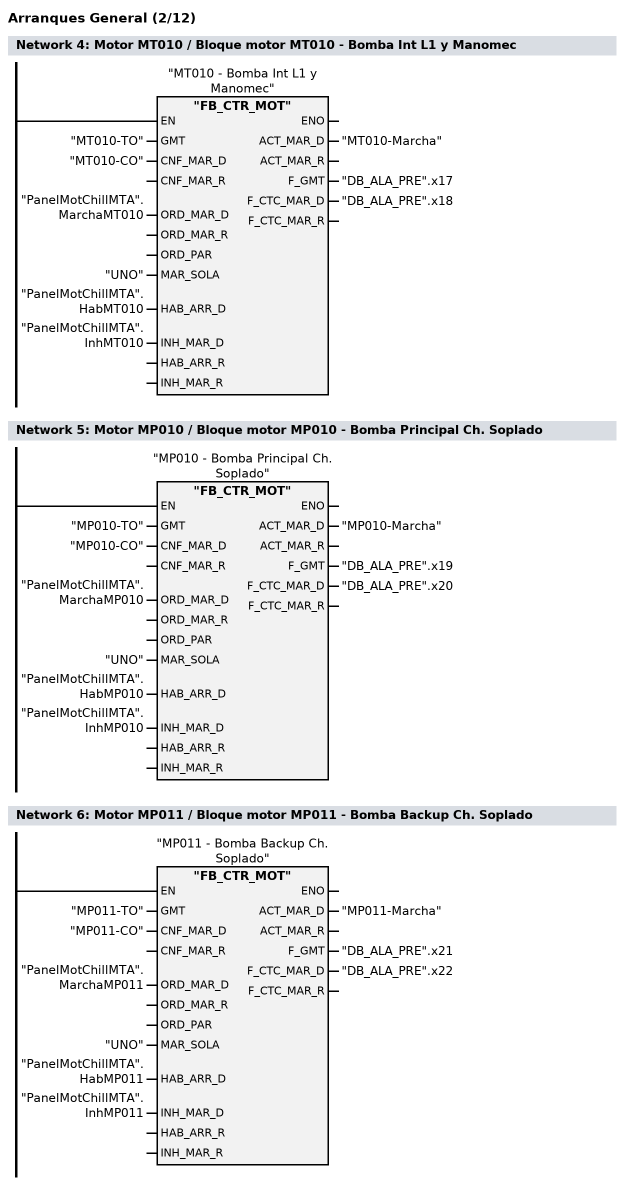
   RUNG wire#powerrail
      "MT010 - Bomba Int L1 y Manomec"(GMT := "MT010-TO", CNF_MAR_D := "MT010-CO", CNF_MAR_R :=, ORD_MAR_D := "PanelMotChillMTA".MarchaMT010, ORD_MAR_R :=, ORD_PAR :=, MAR_SOLA := "UNO", HAB_ARR_D := "PanelMotChillMTA".HabMT010, INH_MAR_D := "PanelMotChillMTA".InhMT010, HAB_ARR_R :=, INH_MAR_R :=, ACT_MAR_D => "MT010-Marcha", ACT_MAR_R =>, F_GMT => "DB_ALA_PRE".x17, F_CTC_MAR_D => "DB_ALA_PRE".x18, F_CTC_MAR_R =>)
   END_RUNG
   // the same network as SCL:
   "MT010 - Bomba Int L1 y Manomec"(GMT := "MT010-TO",   // "FB_CTR_MOT"
                           CNF_MAR_D := "MT010-CO",
                           ORD_MAR_D := "PanelMotChillMTA".MarchaMT010,
                           MAR_SOLA := "UNO",
                           HAB_ARR_D := "PanelMotChillMTA".HabMT010,
                           INH_MAR_D := "PanelMotChillMTA".InhMT010,
                           ACT_MAR_D => "MT010-Marcha",
                           F_GMT => "DB_ALA_PRE".x17,
                           F_CTC_MAR_D => "DB_ALA_PRE".x18);
END_REGION

REGION Network 5: Motor MP010 / Bloque motor MP010 - Bomba Principal Ch. Soplado
   RUNG wire#powerrail
      "MP010 - Bomba Principal Ch. Soplado"(GMT := "MP010-TO", CNF_MAR_D := "MP010-CO", CNF_MAR_R :=, ORD_MAR_D := "PanelMotChillMTA".MarchaMP010, ORD_MAR_R :=, ORD_PAR :=, MAR_SOLA := "UNO", HAB_ARR_D := "PanelMotChillMTA".HabMP010, INH_MAR_D := "PanelMotChillMTA".InhMP010, HAB_ARR_R :=, INH_MAR_R :=, ACT_MAR_D => "MP010-Marcha", ACT_MAR_R =>, F_GMT => "DB_ALA_PRE".x19, F_CTC_MAR_D => "DB_ALA_PRE".x20, F_CTC_MAR_R =>)
   END_RUNG
   // the same network as SCL:
   "MP010 - Bomba Principal Ch. Soplado"(GMT := "MP010-TO",   // "FB_CTR_MOT"
                           CNF_MAR_D := "MP010-CO",
                           ORD_MAR_D := "PanelMotChillMTA".MarchaMP010,
                           MAR_SOLA := "UNO",
                           HAB_ARR_D := "PanelMotChillMTA".HabMP010,
                           INH_MAR_D := "PanelMotChillMTA".InhMP010,
                           ACT_MAR_D => "MP010-Marcha",
                           F_GMT => "DB_ALA_PRE".x19,
                           F_CTC_MAR_D => "DB_ALA_PRE".x20);
END_REGION

REGION Network 6: Motor MP011 / Bloque motor MP011 - Bomba Backup Ch. Soplado
   RUNG wire#powerrail
      "MP011 - Bomba Backup Ch. Soplado"(GMT := "MP011-TO", CNF_MAR_D := "MP011-CO", CNF_MAR_R :=, ORD_MAR_D := "PanelMotChillMTA".MarchaMP011, ORD_MAR_R :=, ORD_PAR :=, MAR_SOLA := "UNO", HAB_ARR_D := "PanelMotChillMTA".HabMP011, INH_MAR_D := "PanelMotChillMTA".InhMP011, HAB_ARR_R :=, INH_MAR_R :=, ACT_MAR_D => "MP011-Marcha", ACT_MAR_R =>, F_GMT => "DB_ALA_PRE".x21, F_CTC_MAR_D => "DB_ALA_PRE".x22, F_CTC_MAR_R =>)
   END_RUNG
   // the same network as SCL:
   "MP011 - Bomba Backup Ch. Soplado"(GMT := "MP011-TO",   // "FB_CTR_MOT"
                           CNF_MAR_D := "MP011-CO",
                           ORD_MAR_D := "PanelMotChillMTA".MarchaMP011,
                           MAR_SOLA := "UNO",
                           HAB_ARR_D := "PanelMotChillMTA".HabMP011,
                           INH_MAR_D := "PanelMotChillMTA".InhMP011,
                           ACT_MAR_D => "MP011-Marcha",
                           F_GMT => "DB_ALA_PRE".x21,
                           F_CTC_MAR_D => "DB_ALA_PRE".x22);
END_REGION

REGION Network 7: Motor MP012 / Bloque motor MP012 - Bomba Principal Ch. Envasado
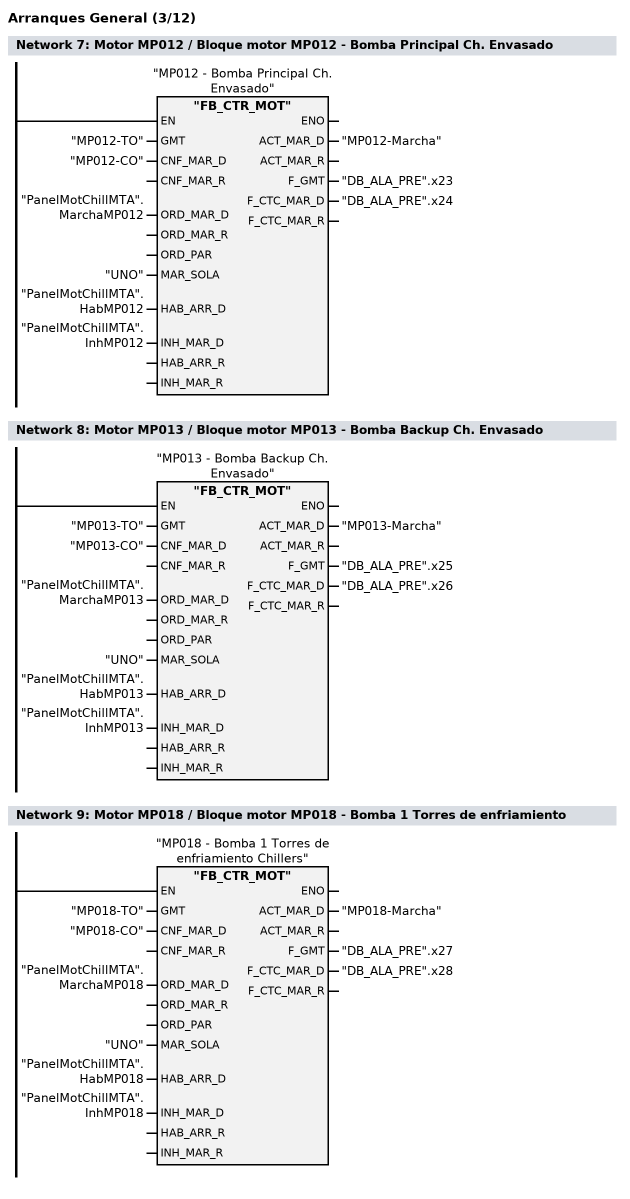
   RUNG wire#powerrail
      "MP012 - Bomba Principal Ch. Envasado"(GMT := "MP012-TO", CNF_MAR_D := "MP012-CO", CNF_MAR_R :=, ORD_MAR_D := "PanelMotChillMTA".MarchaMP012, ORD_MAR_R :=, ORD_PAR :=, MAR_SOLA := "UNO", HAB_ARR_D := "PanelMotChillMTA".HabMP012, INH_MAR_D := "PanelMotChillMTA".InhMP012, HAB_ARR_R :=, INH_MAR_R :=, ACT_MAR_D => "MP012-Marcha", ACT_MAR_R =>, F_GMT => "DB_ALA_PRE".x23, F_CTC_MAR_D => "DB_ALA_PRE".x24, F_CTC_MAR_R =>)
   END_RUNG
   // the same network as SCL:
   "MP012 - Bomba Principal Ch. Envasado"(GMT := "MP012-TO",   // "FB_CTR_MOT"
                           CNF_MAR_D := "MP012-CO",
                           ORD_MAR_D := "PanelMotChillMTA".MarchaMP012,
                           MAR_SOLA := "UNO",
                           HAB_ARR_D := "PanelMotChillMTA".HabMP012,
                           INH_MAR_D := "PanelMotChillMTA".InhMP012,
                           ACT_MAR_D => "MP012-Marcha",
                           F_GMT => "DB_ALA_PRE".x23,
                           F_CTC_MAR_D => "DB_ALA_PRE".x24);
END_REGION

REGION Network 8: Motor MP013 / Bloque motor MP013 - Bomba Backup Ch. Envasado
   RUNG wire#powerrail
      "MP013 - Bomba Backup Ch. Envasado"(GMT := "MP013-TO", CNF_MAR_D := "MP013-CO", CNF_MAR_R :=, ORD_MAR_D := "PanelMotChillMTA".MarchaMP013, ORD_MAR_R :=, ORD_PAR :=, MAR_SOLA := "UNO", HAB_ARR_D := "PanelMotChillMTA".HabMP013, INH_MAR_D := "PanelMotChillMTA".InhMP013, HAB_ARR_R :=, INH_MAR_R :=, ACT_MAR_D => "MP013-Marcha", ACT_MAR_R =>, F_GMT => "DB_ALA_PRE".x25, F_CTC_MAR_D => "DB_ALA_PRE".x26, F_CTC_MAR_R =>)
   END_RUNG
   // the same network as SCL:
   "MP013 - Bomba Backup Ch. Envasado"(GMT := "MP013-TO",   // "FB_CTR_MOT"
                           CNF_MAR_D := "MP013-CO",
                           ORD_MAR_D := "PanelMotChillMTA".MarchaMP013,
                           MAR_SOLA := "UNO",
                           HAB_ARR_D := "PanelMotChillMTA".HabMP013,
                           INH_MAR_D := "PanelMotChillMTA".InhMP013,
                           ACT_MAR_D => "MP013-Marcha",
                           F_GMT => "DB_ALA_PRE".x25,
                           F_CTC_MAR_D => "DB_ALA_PRE".x26);
END_REGION

REGION Network 9: Motor MP018 / Bloque motor MP018 - Bomba 1 Torres de enfriamiento
   RUNG wire#powerrail
      "MP018 - Bomba 1 Torres de enfriamiento Chillers"(GMT := "MP018-TO", CNF_MAR_D := "MP018-CO", CNF_MAR_R :=, ORD_MAR_D := "PanelMotChillMTA".MarchaMP018, ORD_MAR_R :=, ORD_PAR :=, MAR_SOLA := "UNO", HAB_ARR_D := "PanelMotChillMTA".HabMP018, INH_MAR_D := "PanelMotChillMTA".InhMP018, HAB_ARR_R :=, INH_MAR_R :=, ACT_MAR_D => "MP018-Marcha", ACT_MAR_R =>, F_GMT => "DB_ALA_PRE".x27, F_CTC_MAR_D => "DB_ALA_PRE".x28, F_CTC_MAR_R =>)
   END_RUNG
   // the same network as SCL:
   "MP018 - Bomba 1 Torres de enfriamiento Chillers"(GMT := "MP018-TO",   // "FB_CTR_MOT"
                           CNF_MAR_D := "MP018-CO",
                           ORD_MAR_D := "PanelMotChillMTA".MarchaMP018,
                           MAR_SOLA := "UNO",
                           HAB_ARR_D := "PanelMotChillMTA".HabMP018,
                           INH_MAR_D := "PanelMotChillMTA".InhMP018,
                           ACT_MAR_D => "MP018-Marcha",
                           F_GMT => "DB_ALA_PRE".x27,
                           F_CTC_MAR_D => "DB_ALA_PRE".x28);
END_REGION

REGION Network 10: Motor MP019 / Bloque motor MP019 - Bomba 2 Torres de enfriamiento
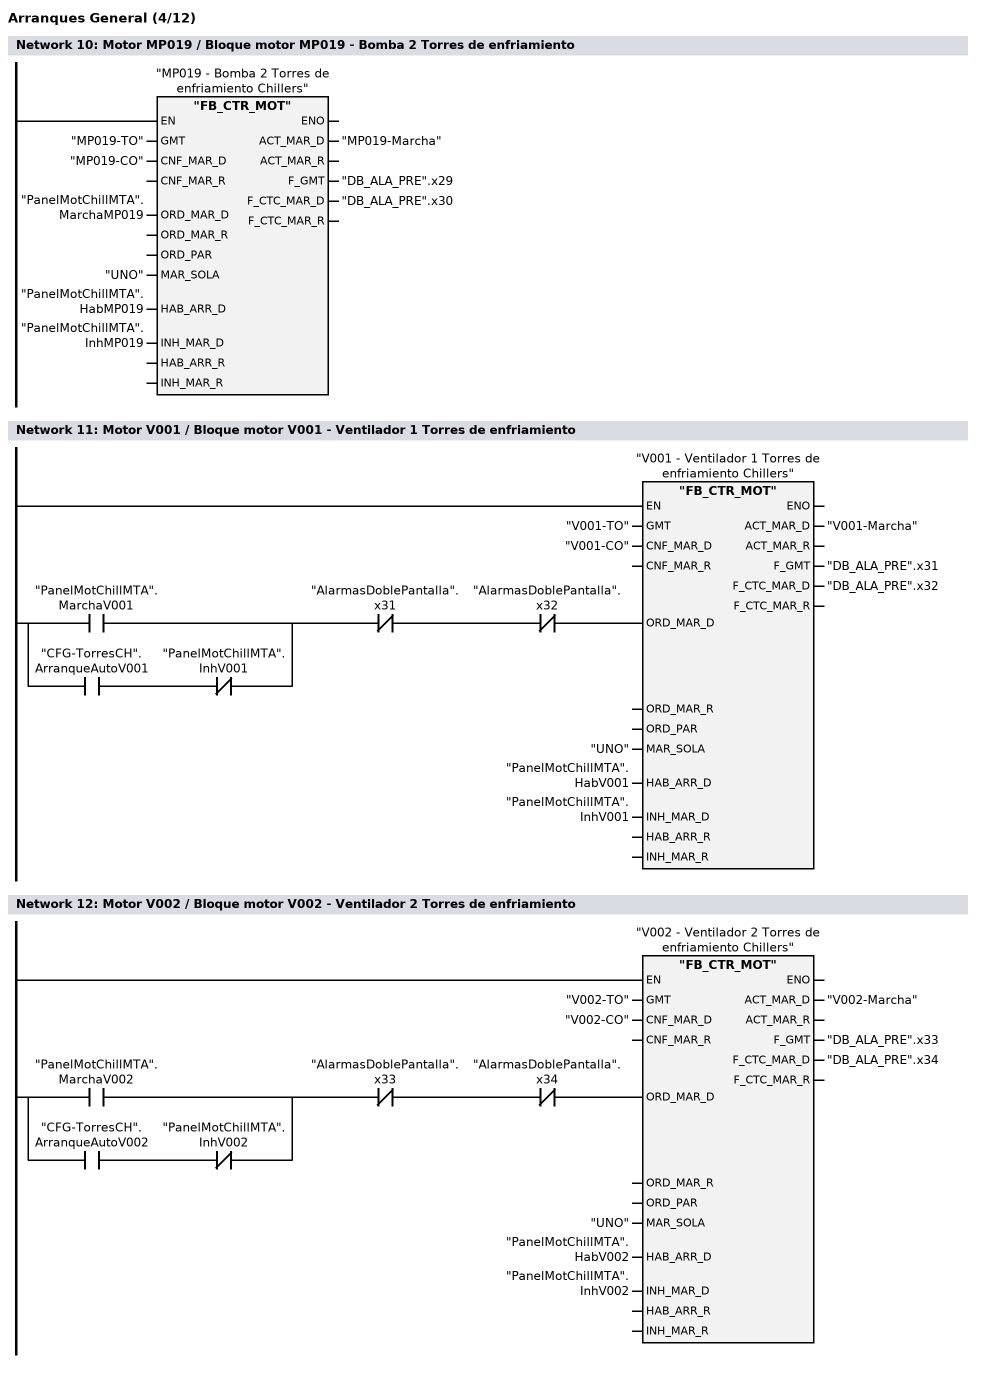
   RUNG wire#powerrail
      "MP019 - Bomba 2 Torres de enfriamiento Chillers"(GMT := "MP019-TO", CNF_MAR_D := "MP019-CO", CNF_MAR_R :=, ORD_MAR_D := "PanelMotChillMTA".MarchaMP019, ORD_MAR_R :=, ORD_PAR :=, MAR_SOLA := "UNO", HAB_ARR_D := "PanelMotChillMTA".HabMP019, INH_MAR_D := "PanelMotChillMTA".InhMP019, HAB_ARR_R :=, INH_MAR_R :=, ACT_MAR_D => "MP019-Marcha", ACT_MAR_R =>, F_GMT => "DB_ALA_PRE".x29, F_CTC_MAR_D => "DB_ALA_PRE".x30, F_CTC_MAR_R =>)
   END_RUNG
   // the same network as SCL:
   "MP019 - Bomba 2 Torres de enfriamiento Chillers"(GMT := "MP019-TO",   // "FB_CTR_MOT"
                           CNF_MAR_D := "MP019-CO",
                           ORD_MAR_D := "PanelMotChillMTA".MarchaMP019,
                           MAR_SOLA := "UNO",
                           HAB_ARR_D := "PanelMotChillMTA".HabMP019,
                           INH_MAR_D := "PanelMotChillMTA".InhMP019,
                           ACT_MAR_D => "MP019-Marcha",
                           F_GMT => "DB_ALA_PRE".x29,
                           F_CTC_MAR_D => "DB_ALA_PRE".x30);
END_REGION

REGION Network 11: Motor V001 / Bloque motor V001 - Ventilador 1 Torres de enfriamiento
   RUNG wire#powerrail
      "V001 - Ventilador 1 Torres de enfriamiento Chillers"(ORD_MAR_D := wire#w2, GMT := "V001-TO", CNF_MAR_D := "V001-CO", CNF_MAR_R :=, ORD_MAR_R :=, ORD_PAR :=, MAR_SOLA := "UNO", HAB_ARR_D := "PanelMotChillMTA".HabV001, INH_MAR_D := "PanelMotChillMTA".InhV001, HAB_ARR_R :=, INH_MAR_R :=, ACT_MAR_D => "V001-Marcha", ACT_MAR_R =>, F_GMT => "DB_ALA_PRE".x31, F_CTC_MAR_D => "DB_ALA_PRE".x32, F_CTC_MAR_R =>)
   END_RUNG
   RUNG wire#powerrail
      Contact( "PanelMotChillMTA".MarchaV001 )
      wire#w1
      I_Contact( "AlarmasDoblePantalla".x31 )
      I_Contact( "AlarmasDoblePantalla".x32 )
   END_RUNG wire#w2
   RUNG wire#powerrail
      Contact( "CFG-TorresCH".ArranqueAutoV001 )
      I_Contact( "PanelMotChillMTA".InhV001 )
   END_RUNG wire#w1
   // the same network as SCL:
   "V001 - Ventilador 1 Torres de enfriamiento Chillers"(GMT := "V001-TO",   // "FB_CTR_MOT"
                           CNF_MAR_D := "V001-CO",
                           ORD_MAR_D := ("PanelMotChillMTA".MarchaV001 OR ("CFG-TorresCH".ArranqueAutoV001 AND NOT "PanelMotChillMTA".InhV001)) AND NOT "AlarmasDoblePantalla".x31 AND NOT "AlarmasDoblePantalla".x32,
                           MAR_SOLA := "UNO",
                           HAB_ARR_D := "PanelMotChillMTA".HabV001,
                           INH_MAR_D := "PanelMotChillMTA".InhV001,
                           ACT_MAR_D => "V001-Marcha",
                           F_GMT => "DB_ALA_PRE".x31,
                           F_CTC_MAR_D => "DB_ALA_PRE".x32);
END_REGION

REGION Network 12: Motor V002 / Bloque motor V002 - Ventilador 2 Torres de enfriamiento
   RUNG wire#powerrail
      "V002 - Ventilador 2 Torres de enfriamiento Chillers"(ORD_MAR_D := wire#w2, GMT := "V002-TO", CNF_MAR_D := "V002-CO", CNF_MAR_R :=, ORD_MAR_R :=, ORD_PAR :=, MAR_SOLA := "UNO", HAB_ARR_D := "PanelMotChillMTA".HabV002, INH_MAR_D := "PanelMotChillMTA".InhV002, HAB_ARR_R :=, INH_MAR_R :=, ACT_MAR_D => "V002-Marcha", ACT_MAR_R =>, F_GMT => "DB_ALA_PRE".x33, F_CTC_MAR_D => "DB_ALA_PRE".x34, F_CTC_MAR_R =>)
   END_RUNG
   RUNG wire#powerrail
      Contact( "PanelMotChillMTA".MarchaV002 )
      wire#w1
      I_Contact( "AlarmasDoblePantalla".x33 )
      I_Contact( "AlarmasDoblePantalla".x34 )
   END_RUNG wire#w2
   RUNG wire#powerrail
      Contact( "CFG-TorresCH".ArranqueAutoV002 )
      I_Contact( "PanelMotChillMTA".InhV002 )
   END_RUNG wire#w1
   // the same network as SCL:
   "V002 - Ventilador 2 Torres de enfriamiento Chillers"(GMT := "V002-TO",   // "FB_CTR_MOT"
                           CNF_MAR_D := "V002-CO",
                           ORD_MAR_D := ("PanelMotChillMTA".MarchaV002 OR ("CFG-TorresCH".ArranqueAutoV002 AND NOT "PanelMotChillMTA".InhV002)) AND NOT "AlarmasDoblePantalla".x33 AND NOT "AlarmasDoblePantalla".x34,
                           MAR_SOLA := "UNO",
                           HAB_ARR_D := "PanelMotChillMTA".HabV002,
                           INH_MAR_D := "PanelMotChillMTA".InhV002,
                           ACT_MAR_D => "V002-Marcha",
                           F_GMT => "DB_ALA_PRE".x33,
                           F_CTC_MAR_D => "DB_ALA_PRE".x34);
END_REGION

REGION Network 13: Motor V003 / Bloque motor V003 - Ventilador 3 Torres de enfriamiento
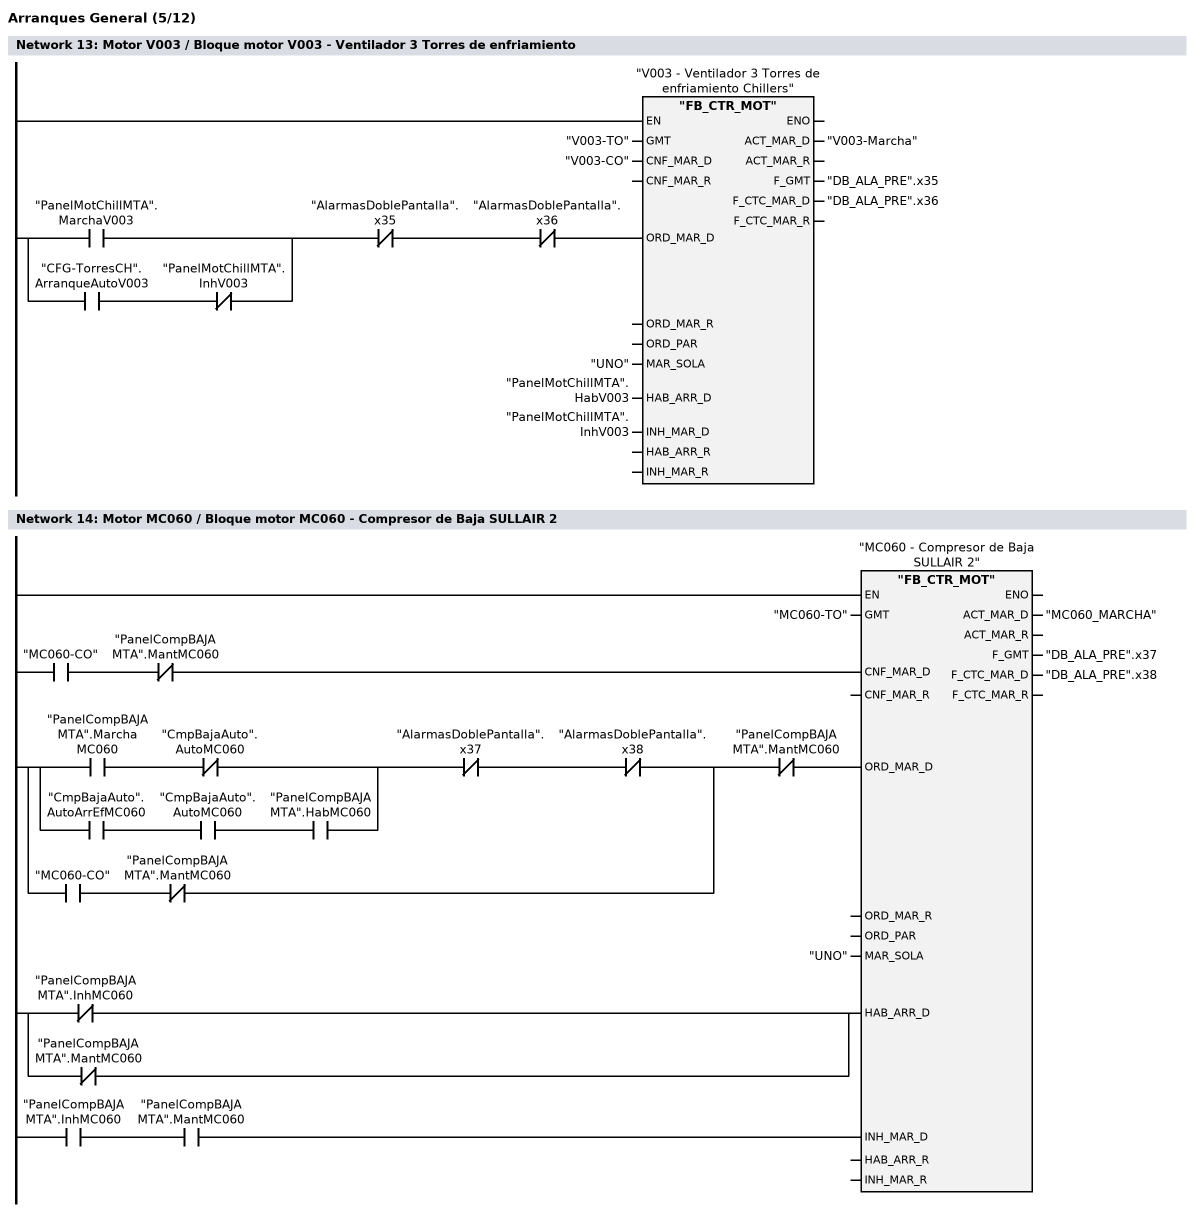
   RUNG wire#powerrail
      "V003 - Ventilador 3 Torres de enfriamiento Chillers"(ORD_MAR_D := wire#w2, GMT := "V003-TO", CNF_MAR_D := "V003-CO", CNF_MAR_R :=, ORD_MAR_R :=, ORD_PAR :=, MAR_SOLA := "UNO", HAB_ARR_D := "PanelMotChillMTA".HabV003, INH_MAR_D := "PanelMotChillMTA".InhV003, HAB_ARR_R :=, INH_MAR_R :=, ACT_MAR_D => "V003-Marcha", ACT_MAR_R =>, F_GMT => "DB_ALA_PRE".x35, F_CTC_MAR_D => "DB_ALA_PRE".x36, F_CTC_MAR_R =>)
   END_RUNG
   RUNG wire#powerrail
      Contact( "PanelMotChillMTA".MarchaV003 )
      wire#w1
      I_Contact( "AlarmasDoblePantalla".x35 )
      I_Contact( "AlarmasDoblePantalla".x36 )
   END_RUNG wire#w2
   RUNG wire#powerrail
      Contact( "CFG-TorresCH".ArranqueAutoV003 )
      I_Contact( "PanelMotChillMTA".InhV003 )
   END_RUNG wire#w1
   // the same network as SCL:
   "V003 - Ventilador 3 Torres de enfriamiento Chillers"(GMT := "V003-TO",   // "FB_CTR_MOT"
                           CNF_MAR_D := "V003-CO",
                           ORD_MAR_D := ("PanelMotChillMTA".MarchaV003 OR ("CFG-TorresCH".ArranqueAutoV003 AND NOT "PanelMotChillMTA".InhV003)) AND NOT "AlarmasDoblePantalla".x35 AND NOT "AlarmasDoblePantalla".x36,
                           MAR_SOLA := "UNO",
                           HAB_ARR_D := "PanelMotChillMTA".HabV003,
                           INH_MAR_D := "PanelMotChillMTA".InhV003,
                           ACT_MAR_D => "V003-Marcha",
                           F_GMT => "DB_ALA_PRE".x35,
                           F_CTC_MAR_D => "DB_ALA_PRE".x36);
END_REGION

REGION Network 14: Motor MC060 / Bloque motor MC060 - Compresor de Baja SULLAIR 2
   RUNG wire#powerrail
      "MC060 - Compresor de Baja SULLAIR 2"(CNF_MAR_D := wire#w1, ORD_MAR_D := wire#w4, HAB_ARR_D := wire#w5, INH_MAR_D := wire#w6, GMT := "MC060-TO", CNF_MAR_R :=, ORD_MAR_R :=, ORD_PAR :=, MAR_SOLA := "UNO", HAB_ARR_R :=, INH_MAR_R :=, ACT_MAR_D => "MC060_MARCHA", ACT_MAR_R =>, F_GMT => "DB_ALA_PRE".x37, F_CTC_MAR_D => "DB_ALA_PRE".x38, F_CTC_MAR_R =>)
   END_RUNG
   RUNG wire#powerrail
      Contact( "MC060-CO" )
      I_Contact( "PanelCompBAJA MTA".MantMC060 )
   END_RUNG wire#w1
   RUNG wire#powerrail
      Contact( "PanelCompBAJA MTA".MarchaMC060 )
      I_Contact( "CmpBajaAuto".AutoMC060 )
      wire#w2
      I_Contact( "AlarmasDoblePantalla".x37 )
      I_Contact( "AlarmasDoblePantalla".x38 )
      wire#w3
      I_Contact( "PanelCompBAJA MTA".MantMC060 )
   END_RUNG wire#w4
   RUNG wire#powerrail
      Contact( "CmpBajaAuto".AutoArrEfMC060 )
      Contact( "CmpBajaAuto".AutoMC060 )
      Contact( "PanelCompBAJA MTA".HabMC060 )
   END_RUNG wire#w2
   RUNG wire#powerrail
      Contact( "MC060-CO" )
      I_Contact( "PanelCompBAJA MTA".MantMC060 )
   END_RUNG wire#w3
   RUNG wire#powerrail
      I_Contact( "PanelCompBAJA MTA".InhMC060 )
   END_RUNG wire#w5
   RUNG wire#powerrail
      I_Contact( "PanelCompBAJA MTA".MantMC060 )
   END_RUNG wire#w5
   RUNG wire#powerrail
      Contact( "PanelCompBAJA MTA".InhMC060 )
      Contact( "PanelCompBAJA MTA".MantMC060 )
   END_RUNG wire#w6
   // the same network as SCL:
   "MC060 - Compresor de Baja SULLAIR 2"(GMT := "MC060-TO",   // "FB_CTR_MOT"
                           CNF_MAR_D := "MC060-CO" AND NOT "PanelCompBAJA MTA".MantMC060,
                           ORD_MAR_D := (((("PanelCompBAJA MTA".MarchaMC060 AND NOT "CmpBajaAuto".AutoMC060) OR ("CmpBajaAuto".AutoArrEfMC060 AND "CmpBajaAuto".AutoMC060 AND "PanelCompBAJA MTA".HabMC060)) AND NOT "AlarmasDoblePantalla".x37 AND NOT "AlarmasDoblePantalla".x38) OR ("MC060-CO" AND NOT "PanelCompBAJA MTA".MantMC060)) AND NOT "PanelCompBAJA MTA".MantMC060,
                           MAR_SOLA := "UNO",
                           HAB_ARR_D := NOT "PanelCompBAJA MTA".InhMC060 OR NOT "PanelCompBAJA MTA".MantMC060,
                           INH_MAR_D := "PanelCompBAJA MTA".InhMC060 AND "PanelCompBAJA MTA".MantMC060,
                           ACT_MAR_D => "MC060_MARCHA",
                           F_GMT => "DB_ALA_PRE".x37,
                           F_CTC_MAR_D => "DB_ALA_PRE".x38);
END_REGION

REGION Network 15
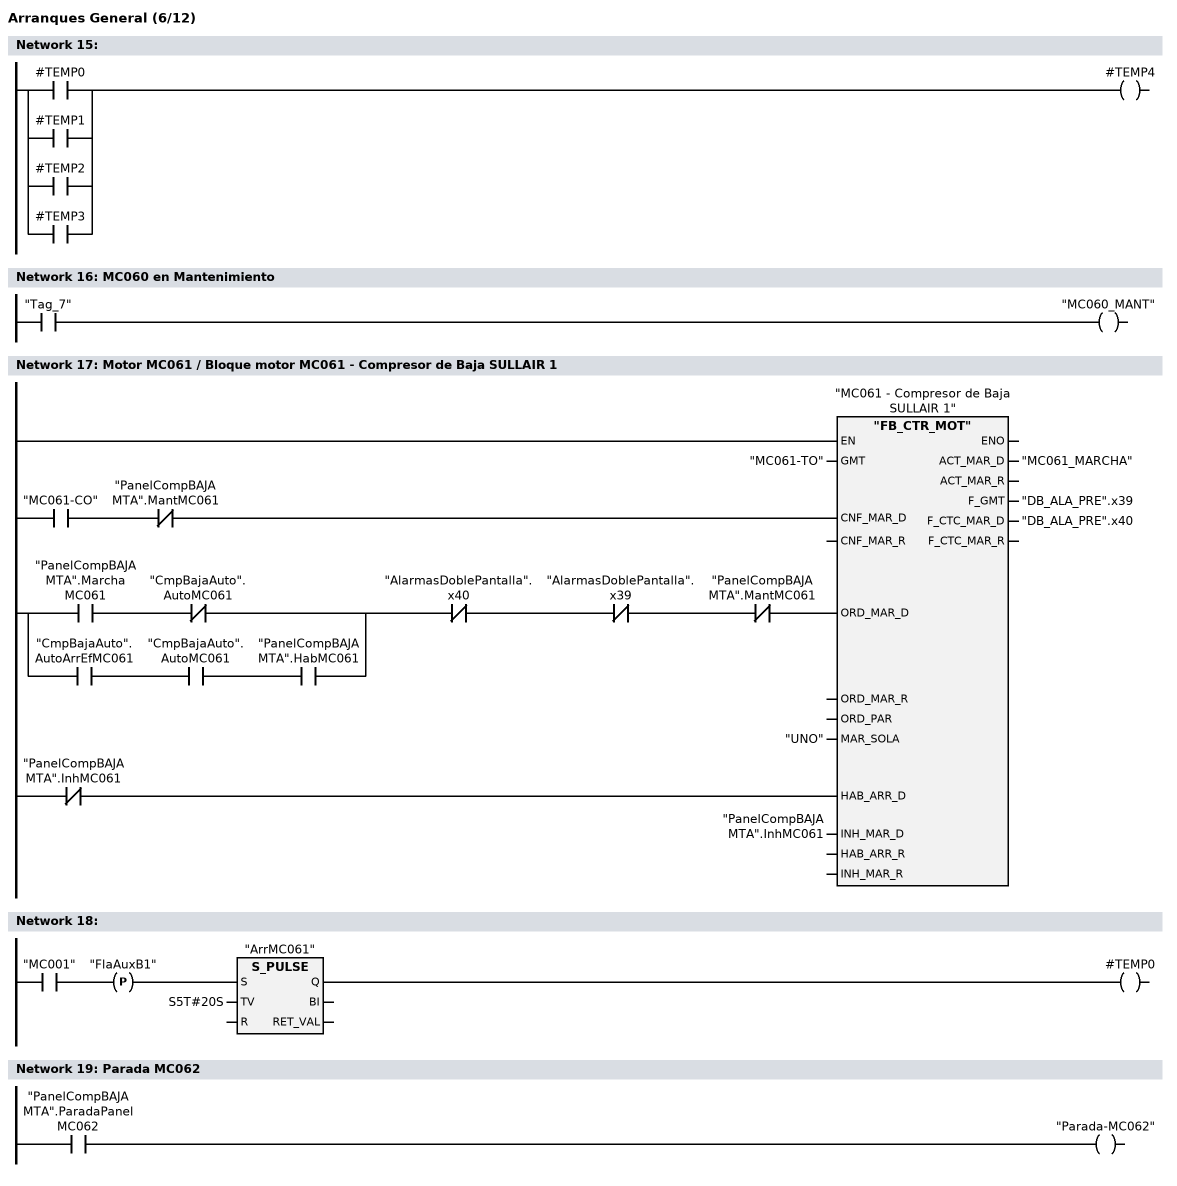
   RUNG wire#powerrail
      Contact( #TEMP0 )
      wire#w1
      Coil( #TEMP4 )
   END_RUNG
   RUNG wire#powerrail
      Contact( #TEMP1 )
   END_RUNG wire#w1
   RUNG wire#powerrail
      Contact( #TEMP2 )
   END_RUNG wire#w1
   RUNG wire#powerrail
      Contact( #TEMP3 )
   END_RUNG wire#w1
   // the same network as SCL:
   #TEMP4 := #TEMP0 OR #TEMP1 OR #TEMP2 OR #TEMP3;
END_REGION

REGION Network 16: MC060 en Mantenimiento
   RUNG wire#powerrail
      Contact( "Tag_7" )
      Coil( "MC060_MANT" )
   END_RUNG
   // the same network as SCL:
   "MC060_MANT" := "Tag_7";
END_REGION

REGION Network 17: Motor MC061 / Bloque motor MC061 - Compresor de Baja SULLAIR 1
   RUNG wire#powerrail
      "MC061 - Compresor de Baja SULLAIR 1"(CNF_MAR_D := wire#w1, ORD_MAR_D := wire#w3, HAB_ARR_D := wire#w4, GMT := "MC061-TO", CNF_MAR_R :=, ORD_MAR_R :=, ORD_PAR :=, MAR_SOLA := "UNO", INH_MAR_D := "PanelCompBAJA MTA".InhMC061, HAB_ARR_R :=, INH_MAR_R :=, ACT_MAR_D => "MC061_MARCHA", ACT_MAR_R =>, F_GMT => "DB_ALA_PRE".x39, F_CTC_MAR_D => "DB_ALA_PRE".x40, F_CTC_MAR_R =>)
   END_RUNG
   RUNG wire#powerrail
      Contact( "MC061-CO" )
      I_Contact( "PanelCompBAJA MTA".MantMC061 )
   END_RUNG wire#w1
   RUNG wire#powerrail
      Contact( "PanelCompBAJA MTA".MarchaMC061 )
      I_Contact( "CmpBajaAuto".AutoMC061 )
      wire#w2
      I_Contact( "AlarmasDoblePantalla".x40 )
      I_Contact( "AlarmasDoblePantalla".x39 )
      I_Contact( "PanelCompBAJA MTA".MantMC061 )
   END_RUNG wire#w3
   RUNG wire#powerrail
      Contact( "CmpBajaAuto".AutoArrEfMC061 )
      Contact( "CmpBajaAuto".AutoMC061 )
      Contact( "PanelCompBAJA MTA".HabMC061 )
   END_RUNG wire#w2
   RUNG wire#powerrail
      I_Contact( "PanelCompBAJA MTA".InhMC061 )
   END_RUNG wire#w4
   // the same network as SCL:
   "MC061 - Compresor de Baja SULLAIR 1"(GMT := "MC061-TO",   // "FB_CTR_MOT"
                           CNF_MAR_D := "MC061-CO" AND NOT "PanelCompBAJA MTA".MantMC061,
                           ORD_MAR_D := (("PanelCompBAJA MTA".MarchaMC061 AND NOT "CmpBajaAuto".AutoMC061) OR ("CmpBajaAuto".AutoArrEfMC061 AND "CmpBajaAuto".AutoMC061 AND "PanelCompBAJA MTA".HabMC061)) AND NOT "AlarmasDoblePantalla".x40 AND NOT "AlarmasDoblePantalla".x39 AND NOT "PanelCompBAJA MTA".MantMC061,
                           MAR_SOLA := "UNO",
                           HAB_ARR_D := NOT "PanelCompBAJA MTA".InhMC061,
                           INH_MAR_D := "PanelCompBAJA MTA".InhMC061,
                           ACT_MAR_D => "MC061_MARCHA",
                           F_GMT => "DB_ALA_PRE".x39,
                           F_CTC_MAR_D => "DB_ALA_PRE".x40);
END_REGION

REGION Network 18
   RUNG wire#powerrail
      Contact( "MC001" )
      P_Trig( "FlaAuxB1" )
      S_PULSE(T_NO := "ArrMC061", TV := S5T#20S, R :=, BI =>, RET_VAL =>)
      Coil( #TEMP0 )
   END_RUNG
   // the same network as SCL:
   #_w1 := "MC001" AND NOT "FlaAuxB1";   // rising edge
   "FlaAuxB1" := "MC001";
   #_s5time1 := S_PULSE(T_NO := "ArrMC061", S := #_w1, TV := S5T#20S, Q => #_w2);
   #TEMP0 := #_w2;
END_REGION

REGION Network 19: Parada MC062
   RUNG wire#powerrail
      Contact( "PanelCompBAJA MTA".ParadaPanelMC062 )
      Coil( "Parada-MC062" )
   END_RUNG
   // the same network as SCL:
   "Parada-MC062" := "PanelCompBAJA MTA".ParadaPanelMC062;
END_REGION

REGION Network 20: Motor MC062 / Bloque motor MC062 - Compresor de Baja SULLAIR 0
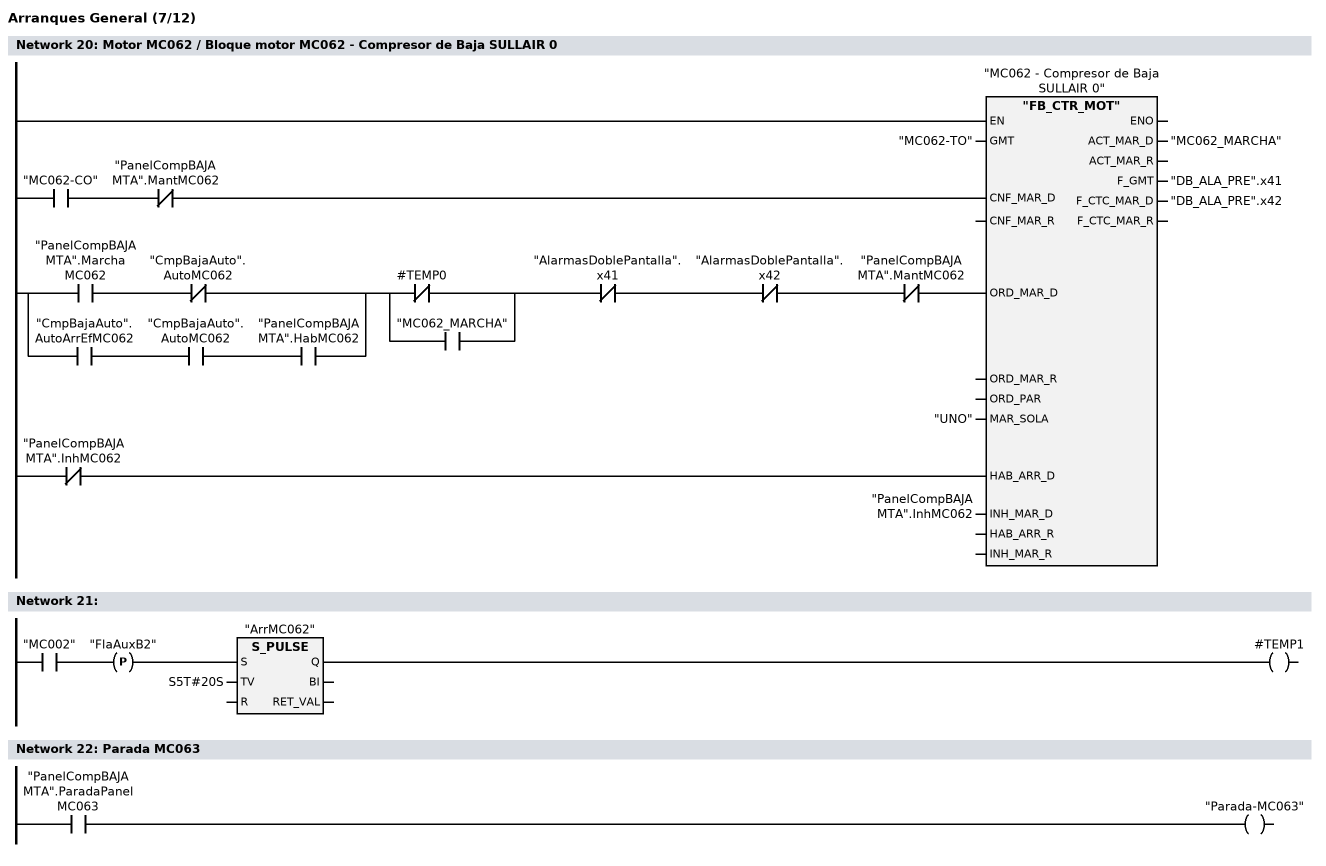
   RUNG wire#powerrail
      "MC062 - Compresor de Baja SULLAIR 0"(CNF_MAR_D := wire#w1, ORD_MAR_D := wire#w4, HAB_ARR_D := wire#w5, GMT := "MC062-TO", CNF_MAR_R :=, ORD_MAR_R :=, ORD_PAR :=, MAR_SOLA := "UNO", INH_MAR_D := "PanelCompBAJA MTA".InhMC062, HAB_ARR_R :=, INH_MAR_R :=, ACT_MAR_D => "MC062_MARCHA", ACT_MAR_R =>, F_GMT => "DB_ALA_PRE".x41, F_CTC_MAR_D => "DB_ALA_PRE".x42, F_CTC_MAR_R =>)
   END_RUNG
   RUNG wire#powerrail
      Contact( "MC062-CO" )
      I_Contact( "PanelCompBAJA MTA".MantMC062 )
   END_RUNG wire#w1
   RUNG wire#powerrail
      Contact( "PanelCompBAJA MTA".MarchaMC062 )
      I_Contact( "CmpBajaAuto".AutoMC062 )
      wire#w2
      I_Contact( #TEMP0 )
      wire#w3
      I_Contact( "AlarmasDoblePantalla".x41 )
      I_Contact( "AlarmasDoblePantalla".x42 )
      I_Contact( "PanelCompBAJA MTA".MantMC062 )
   END_RUNG wire#w4
   RUNG wire#powerrail
      Contact( "CmpBajaAuto".AutoArrEfMC062 )
      Contact( "CmpBajaAuto".AutoMC062 )
      Contact( "PanelCompBAJA MTA".HabMC062 )
   END_RUNG wire#w2
   RUNG wire#w2
      Contact( "MC062_MARCHA" )
   END_RUNG wire#w3
   RUNG wire#powerrail
      I_Contact( "PanelCompBAJA MTA".InhMC062 )
   END_RUNG wire#w5
   // the same network as SCL:
   "MC062 - Compresor de Baja SULLAIR 0"(GMT := "MC062-TO",   // "FB_CTR_MOT"
                           CNF_MAR_D := "MC062-CO" AND NOT "PanelCompBAJA MTA".MantMC062,
                           ORD_MAR_D := (("PanelCompBAJA MTA".MarchaMC062 AND NOT "CmpBajaAuto".AutoMC062) OR ("CmpBajaAuto".AutoArrEfMC062 AND "CmpBajaAuto".AutoMC062 AND "PanelCompBAJA MTA".HabMC062)) AND (NOT #TEMP0 OR "MC062_MARCHA") AND NOT "AlarmasDoblePantalla".x41 AND NOT "AlarmasDoblePantalla".x42 AND NOT "PanelCompBAJA MTA".MantMC062,
                           MAR_SOLA := "UNO",
                           HAB_ARR_D := NOT "PanelCompBAJA MTA".InhMC062,
                           INH_MAR_D := "PanelCompBAJA MTA".InhMC062,
                           ACT_MAR_D => "MC062_MARCHA",
                           F_GMT => "DB_ALA_PRE".x41,
                           F_CTC_MAR_D => "DB_ALA_PRE".x42);
END_REGION

REGION Network 21
   RUNG wire#powerrail
      Contact( "MC002" )
      P_Trig( "FlaAuxB2" )
      S_PULSE(T_NO := "ArrMC062", TV := S5T#20S, R :=, BI =>, RET_VAL =>)
      Coil( #TEMP1 )
   END_RUNG
   // the same network as SCL:
   #_w1 := "MC002" AND NOT "FlaAuxB2";   // rising edge
   "FlaAuxB2" := "MC002";
   #_s5time1 := S_PULSE(T_NO := "ArrMC062", S := #_w1, TV := S5T#20S, Q => #_w2);
   #TEMP1 := #_w2;
END_REGION

REGION Network 22: Parada MC063
   RUNG wire#powerrail
      Contact( "PanelCompBAJA MTA".ParadaPanelMC063 )
      Coil( "Parada-MC063" )
   END_RUNG
   // the same network as SCL:
   "Parada-MC063" := "PanelCompBAJA MTA".ParadaPanelMC063;
END_REGION

REGION Network 23: Motor MC063 / Bloque motor MC063 - Compresor de Baja ATLAS 3